// TIA Portal project "Buffer Station" (V20)
// Programming buffer station with Factory I/O

(* hardware
DEVICE "S7-1200 station_1"  S7-1200 Station
   slot 0: "Rack_0"  S7-1200 Rack  Rack  V1.0
   slot 1: "PLC_1"  CPU 1212C AC/DC/Rly  6ES7 212-1BE40-0XB0  V4.6
DEVICE "HMI_1"  KTP700 Basic PN
   slot 0: "HMI_1"  KTP700 Basic PN  6AV2 123-2GB03-0AX0  17.0.0.0
   slot 1: "HMI_RT_1"  KTP700 Basic PN  6AV2 123-2GB03-0AX0  17.0.0.0
   slot 5: "HMI_1.IE_CP_1"  PROFINET Interface  17.0.0.0
      slot 1: "PROFINET Interface_1"  PROFINET Interface
         slot 1: "Port_1"  Port
*)

// ===== PLC "PLC_1"  CPU 1212C AC/DC/Rly =====

VAR_GLOBAL   // PLC tag table "Inputs"
   "atBufferEntry" AT %I1.0 : Bool;
   "atBufferExit" AT %I1.1 : Bool;
   "atExit" AT %I1.2 : Bool;
   "startButton" AT %I1.3 : Bool;
   "resetButton" AT %I1.4 : Bool;
   "stopButton" AT %I1.5 : Bool;
   "autoMode" AT %I1.6 : Bool;
   "emergencyStop" AT %I1.7 : Bool;
   "bufferVel" AT %ID100 : Real;
   "exitVel" AT %ID104 : Real;
   "Tag_1" AT %MD100 : DWord;
END_VAR

VAR_GLOBAL   // PLC tag table "Outputs"
   "stopBlade" AT %Q0.0 : Bool;
   "startLight" AT %Q0.1 : Bool;
   "resetLight" AT %Q0.2 : Bool;
   "stopLight" AT %Q0.3 : Bool;
   "bufferConveyor" AT %QD100 : Real;
   "exitConveyor" AT %QD104 : Real;
   "counterBoxes" AT %QD108 : DInt;
END_VAR

DATA_BLOCK "Data"   // DB1
{ S7_Optimized_Access := 'TRUE' }
VERSION : 0.1
   VAR
      S_R_Conveyors : Bool := false;   // latch or unlatch conveyors
      Counter_Box : Struct
         fTrigger : Bool;
         currentCount : DInt;
      END_STRUCT;
      freqBufferConveyor : Struct
         stopBladeState : Bool;
         setBlade : Bool;
         resetBlade : Bool;
      END_STRUCT;
      HMI : Struct
         startButton : Bool;
         stopButton : Bool;
         resetButton : Bool;
      END_STRUCT;
   END_VAR
BEGIN
END_DATA_BLOCK

FUNCTION "Start_Stop" : Void   // FC1, SCL
{ S7_Optimized_Access := 'TRUE' }
VERSION : 0.1
   VAR_INPUT
      emergencyStop : Bool;
      stopButton : Bool;
      startButton : Bool;
      resetButton : Bool;
      autoMode : Bool;
      bufferVel : Real;
      exitVel : Real;
      atBufferExit : Bool;
   END_VAR
   VAR_OUTPUT
      bufferConveyor : Real;
      exitConveyor : Real;
      startLight : Bool;
      stopLight : Bool;
   END_VAR
BEGIN
   REGION Conveyors Run
       // RESET All Logic
       IF NOT #emergencyStop OR NOT #stopButton OR NOT #autoMode OR "Data".HMI.stopButton THEN
           "Data".S_R_Conveyors := FALSE;
       END_IF;
       //SET All Logic
       IF #startButton OR "Data".HMI.startButton AND #autoMode THEN
           "Data".S_R_Conveyors := TRUE;
       END_IF;
   END_REGION

   // Indicator Lights Start and Stop
   REGION Indicator Lights
       IF NOT "Data".S_R_Conveyors THEN
           #stopLight := TRUE;
       ELSE
           #startLight := TRUE;
       END_IF;
   END_REGION

   // Control Conveyors
   REGION Frequency Buffer and Exit Conveyor
       IF "Data".S_R_Conveyors THEN
           #exitConveyor := #exitVel;
           #bufferConveyor := #bufferVel;
           IF "Data".freqBufferConveyor.stopBladeState THEN
               #bufferConveyor := 0;
           END_IF;
       END_IF;
   END_REGION
END_FUNCTION

FUNCTION "Counter_Blade_Control" : Void   // FC2, SCL
{ S7_Optimized_Access := 'TRUE' }
VERSION : 0.1
   VAR_INPUT
      atExit : Bool;
      resetCounter : Bool;
      atBufferExit : Bool;
      atBufferEntry : Bool;
   END_VAR
   VAR_OUTPUT
      counterDisplay : DInt;
      resetLight : Bool;
      stopBlade : Bool;
   END_VAR
BEGIN
   // Counter Box Logic
   REGION Box Counter
       // At Exit sensor activate Risind Edge 
       "F_TRIG_COUNT"(CLK:=#atBufferEntry,
                     Q=>"Data".Counter_Box.fTrigger);
      // Reset button gets counter to 0
      IF #resetCounter OR "Data".HMI.resetButton THEN
          "Data".Counter_Box.currentCount := 0;
          #resetLight := TRUE;
          // When the Falling Edge is activated, the count value increase 1
      ELSIF "Data".Counter_Box.fTrigger THEN
          "Data".Counter_Box.currentCount := "Data".Counter_Box.currentCount + 1;
      END_IF;
      #counterDisplay := "Data".Counter_Box.currentCount;
   END_REGION

   // Blade Control Logic
   REGION Blade Control
       IF "Data".S_R_Conveyors THEN
           // At Buffer Exit sensor activate Rising Edge
           "R_TRIG_Blade"(CLK := #atBufferExit,
                          Q => "Data".freqBufferConveyor.setBlade);
           // RESET Blade
           // At Exit sensor reset blade via Rising Edge or if the current counter is less than 2
           "R_TRIG_Exit"(CLK := #atExit,
                         Q => "Data".freqBufferConveyor.resetBlade);
           IF "Data".freqBufferConveyor.resetBlade OR "Data".Counter_Box.currentCount = 0 THEN
               "Data".freqBufferConveyor.stopBladeState := FALSE;
               // SET Blade
           ELSIF "Data".freqBufferConveyor.setBlade THEN
               "Data".freqBufferConveyor.stopBladeState := TRUE;
           END_IF;
       END_IF;
       #stopBlade := "Data".freqBufferConveyor.stopBladeState;
   END_REGION
END_FUNCTION

ORGANIZATION_BLOCK "Main"   // OB1, LAD, ProgramCycle
TITLE = "Main Program Sweep (Cycle)"
{ S7_Optimized_Access := 'TRUE' }
VERSION : 0.1
   VAR_INPUT
      Initial_Call : Bool;   // Initial call of this OB
      Remanence : Bool;   // =True, if remanent data are available
   END_VAR
BEGIN

REGION Network 1
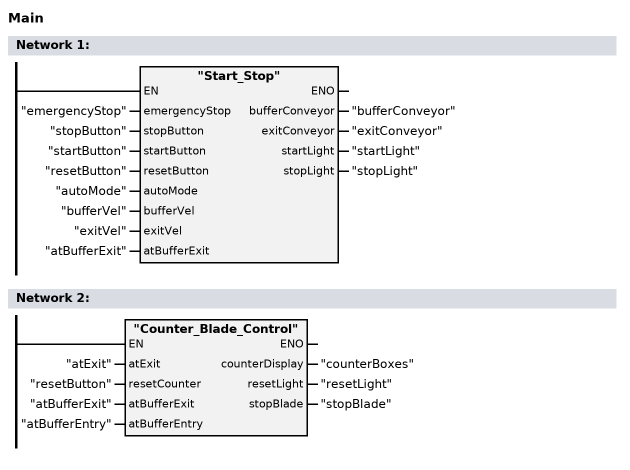
   RUNG wire#powerrail
      "Start_Stop"(emergencyStop := "emergencyStop", stopButton := "stopButton", startButton := "startButton", resetButton := "resetButton", autoMode := "autoMode", bufferVel := "bufferVel", exitVel := "exitVel", atBufferExit := "atBufferExit", bufferConveyor => "bufferConveyor", exitConveyor => "exitConveyor", startLight => "startLight", stopLight => "stopLight")
   END_RUNG
   // the same network as SCL:
   "Start_Stop"(emergencyStop := "emergencyStop",
                stopButton := "stopButton",
                startButton := "startButton",
                resetButton := "resetButton",
                autoMode := "autoMode",
                bufferVel := "bufferVel",
                exitVel := "exitVel",
                atBufferExit := "atBufferExit",
                bufferConveyor => "bufferConveyor",
                exitConveyor => "exitConveyor",
                startLight => "startLight",
                stopLight => "stopLight");
END_REGION

REGION Network 2
   RUNG wire#powerrail
      "Counter_Blade_Control"(atExit := "atExit", resetCounter := "resetButton", atBufferExit := "atBufferExit", atBufferEntry := "atBufferEntry", counterDisplay => "counterBoxes", resetLight => "resetLight", stopBlade => "stopBlade")
   END_RUNG
   // the same network as SCL:
   "Counter_Blade_Control"(atExit := "atExit",
                           resetCounter := "resetButton",
                           atBufferExit := "atBufferExit",
                           atBufferEntry := "atBufferEntry",
                           counterDisplay => "counterBoxes",
                           resetLight => "resetLight",
                           stopBlade => "stopBlade");
END_REGION
END_ORGANIZATION_BLOCK

(* ===== HMI "HMI_RT_1" =====
system functions are stored by id; their names below are inferred from use
connection "HMI_Connection_1": ETHERNET, SMART_S7_1200_OMS

HMI tags "Default tag table"
   "Tag_ScreenNumber" : UInt, internal
   "currentCount" : DInt = PLC Data.Counter_Box.currentCount AT %DB1.DBD0, 100 ms
   "bladeState" : Bool = PLC stopBlade AT %Q0.0, 100 ms
   "atBufferExit" : Bool = PLC atBufferExit AT %I1.1, 100 ms
   "atExit" : Bool = PLC atExit AT %I1.2, 1 s
   "speedBufferConveyor" : Real = PLC bufferConveyor AT %QD100, 100 ms
   "speedExitConveyor" : Real = PLC exitConveyor AT %QD104, 1 s
   "startButton" : Bool = PLC Data.HMI.startButton AT %DB1.DBD0, 1 s
   "stopButton" : Bool = PLC Data.HMI.stopButton AT %DB1.DBD0, 1 s
   "resetButton" : Bool = PLC Data.HMI.resetButton AT %DB1.DBD0, 1 s
   "S_R_State" : Bool = PLC Data.S_R_Conveyors AT %DB1.DBX0.0, 1 s

Template "Template_1" 800x480
   Button "Exit" at 714,429 size 71x50; TextOff 'Exit'; PictureOff "ExitRuntime_KTP700_Basic_PN_TR"; PictureOn "ExitRuntime_KTP700_Basic_PN_TR"
      on Release: StopRuntime(0)
   Button "Template_Button" at 614,429 size 71x50; TextOff 'Text'
   Button "Template_Button_1" at 514,429 size 71x50; TextOff 'Text'
   Button "Template_Button_2" at 414,429 size 71x50; TextOff 'Text'
   Button "Template_Button_3" at 314,429 size 71x50; TextOff 'Text'
   Button "Template_Button_4" at 214,429 size 71x50; TextOff 'Text'
   Button "Alarms" at 114,429 size 71x50; TextOff 'Alarms'; PictureOff "AlarmDisplay_KTP700_Basic_PN_TR"; PictureOn "AlarmDisplay_KTP700_Basic_PN_TR"
      on Release: function_ef3f5d25("Alarm window_Unacknowledged", -1)
   Button "Start screen" at 14,429 size 71x50; TextOff 'Start screen'; PictureOff "NavigateHome_KTP700_Basic_PN_TR"; PictureOn "NavigateHome_KTP700_Basic_PN_TR"
      on Release: ActivateScreen("Root screen", 0)
   SymbolicIOField "Symbolic_IO_Field_Screen" at 187,9 size 506x33; TextOff '0'; TextOn '1'; TextList "TextList_ScreenNames"
      ProcessValue <- "Tag_ScreenNumber"
      on Change: ActivateScreenByNumber("Tag_ScreenNumber", 0)
   DateTimeField "HmiScreenItemData" at 695,25 size 105x25
   DateTimeField "HmiScreenItemData_1" at 695,0 size 105x25
   GraphicView "Logo" at 0,0 size 185x51; Picture "Logo of HMI_1"

screen "Root screen" 800x480, template "Template_1"
   on GenerateScreen: SetTag("Tag_ScreenNumber", 1)
   IOField "I/O field_1" at 120,99 size 132x51; FormatPattern 9999
      ProcessValue <- "currentCount"
   TextField "Text field_1" at 134,68 size 102x23; Text 'Total Boxes'
   Circle "Circle_2" at 504,255 size 28x28
      Appearance <- "bladeState"
   TextField "Text field_3" at 546,258 size 51x23; Text 'Blade'
   Circle "Circle_3" at 504,336 size 28x28
      Appearance <- "atBufferExit"
   TextField "Text field_4" at 546,339 size 116x23; Text 'At Buffer Exit'
   Circle "Circle_4" at 504,377 size 28x28
      Appearance <- "atExit"
   TextField "Text field_5" at 546,380 size 61x23; Text 'At Exit'
   Circle "Circle_1" at 251,321 size 28x28
      Appearance <- "S_R_State"
   TextField "Text field_7" at 531,223 size 76x23; Text 'Actuator'
   TextField "Text field_8" at 532,299 size 68x23; Text 'Sensors'
   Button "Button_1" at 134,175 size 96x32; TextOff 'Reset'
      on Press: function_b14e0dd5("resetButton", 0)
   Button "Button_2" at 134,294 size 96x32; TextOff 'Start'
      on Press: function_b14e0dd5("startButton", 0)
   Button "Button_3" at 134,349 size 96x32; TextOff 'Stop'
      on Press: function_b14e0dd5("stopButton", 0)
   IOField "I/O field_2" at 531,99 size 96x32; FormatPattern 9999
      ProcessValue <- "speedBufferConveyor"
   IOField "I/O field_3" at 531,163 size 96x32; FormatPattern 9999
      ProcessValue <- "speedExitConveyor"
   TextField "Text field_9" at 495,137 size 173x23; Text 'Speed Exit Conveyor'
   TextField "Text field_10" at 495,70 size 191x23; Text 'Speed Buffer Conveyor'
*)